
       FOR #tempLoop := 0 TO #NUM_TYPES DO
           //calculate max # of pages
           #recipeMaxPages[#tempLoop] := DINT_TO_INT(CEIL((#tempSetptsUpper[#tempLoop] - #tempSetptsLower[#tempLoop] + 1.0) / #SETPOINTS_PERPAGE));
           //ensure that current page is within the limits
           #recipeCurrentPages[#tempLoop] := LIMIT(MN := 1, IN := #recipeCurrentPages[#tempLoop], MX := #recipeMaxPages[#tempLoop]);
       END_FOR;

       #recipeMaxPages[4] := DINT_TO_INT(CEIL((#tempNumRecipesUpper - #tempNumRecipesLower + 1.0) / #RECIPES_PERPAGE));
       #recipeCurrentPages[4] := LIMIT(MN := 1, IN := #recipeCurrentPages[4], MX := #recipeMaxPages[4]);
   END_REGION


   REGION REAL
       //index in Setpoints_XXX of the current popup
       #tempCurrentPopup := #recipePopupTrackers[#INDEX_REAL] + #SETPOINTS_PERPAGE * (#recipeCurrentPages[#INDEX_REAL] - 1) + #tempSetptsLower[#INDEX_REAL];

       IF #statPrevPopupTrackers[#INDEX_REAL] <> #recipePopupTrackers[#INDEX_REAL] THEN
           //if a new popup has been loaded, load the new setpoint so they can be displayed
           #recipePopup_REAL := #setpoints_REAL[#tempCurrentPopup];
       ELSE
           //if the HMI popup was updated, relay the commands back to the actual setpoint tag for processing
           //taking care to ensure that changes to the setpoints tags made in other areas of the program do not get overwritten
           IF (#statPrevPopupIN_REAL <> #recipePopup_REAL.IN) AND (#statPrevSetpointIN_REAL = #setpoints_REAL[#tempCurrentPopup].IN) THEN
               #setpoints_REAL[#tempCurrentPopup].IN := #recipePopup_REAL.IN;
           END_IF;
           IF #statPrevPopupsSave[#INDEX_REAL] <> #recipePopup_REAL.SaveSetpoint THEN
               #setpoints_REAL[#tempCurrentPopup].SaveSetpoint := #recipePopup_REAL.SaveSetpoint;
           END_IF;
           IF #statPrevPopupsRevert[#INDEX_REAL] <> #recipePopup_REAL.RevertSetpoint THEN
               #setpoints_REAL[#tempCurrentPopup].RevertSetpoint := #recipePopup_REAL.RevertSetpoint;
           END_IF;

           //then update the popup with the latest setpoint information
           #recipePopup_REAL := #setpoints_REAL[#tempCurrentPopup];
       END_IF;

       //set previous values for next scan
       #statPrevPopupIN_REAL := #recipePopup_REAL.IN;
       #statPrevSetpointIN_REAL := #setpoints_REAL[#tempCurrentPopup].IN;
       #statPrevPopupsSave[#INDEX_REAL] := #recipePopup_REAL.SaveSetpoint;
       #statPrevPopupsRevert[#INDEX_REAL] := #recipePopup_REAL.RevertSetpoint;


       //update main setpoint display with setpoint data
       FOR #tempLoop := 0 TO #SETPOINTS_PERPAGE - 1 DO
           IF #tempLoop + #SETPOINTS_PERPAGE * (#recipeCurrentPages[#INDEX_REAL] - 1) + #tempSetptsLower[#INDEX_REAL] <= #tempSetptsUpper[#INDEX_REAL] THEN
               #setpointsArray_REAL[#tempLoop] := #setpoints_REAL[#tempLoop + #SETPOINTS_PERPAGE * (#recipeCurrentPages[#INDEX_REAL] - 1) + #tempSetptsLower[#INDEX_REAL]];
               #setpointFaceplatesDisable_REAL[#tempLoop] := false;
           ELSE
               #setpointFaceplatesDisable_REAL[#tempLoop] := true;
           END_IF;
       END_FOR;
   END_REGION


   REGION DINT
       //index in Setpoints_XXX of the current popup
       #tempCurrentPopup := #recipePopupTrackers[#INDEX_DINT] + #SETPOINTS_PERPAGE * (#recipeCurrentPages[#INDEX_DINT] - 1) + #tempSetptsLower[#INDEX_DINT];

       IF #statPrevPopupTrackers[#INDEX_DINT] <> #recipePopupTrackers[#INDEX_DINT] THEN
           //if a new popup has been loaded, load the new setpoint so they can be displayed
           #recipePopup_DINT := #setpoints_DINT[#tempCurrentPopup];
       ELSE
           //if the HMI popup was updated, relay the commands back to the actual setpoint tag for processing
           //taking care to ensure that changes to the setpoints tags made in other areas of the program do not get overwritten
           IF (#statPrevPopupIN_DINT <> #recipePopup_DINT.IN) AND (#statPrevSetpointIN_DINT = #setpoints_DINT[#tempCurrentPopup].IN) THEN
               #setpoints_DINT[#tempCurrentPopup].IN := #recipePopup_DINT.IN;
           END_IF;
           IF #statPrevPopupsSave[#INDEX_DINT] <> #recipePopup_DINT.SaveSetpoint THEN
               #setpoints_DINT[#tempCurrentPopup].SaveSetpoint := #recipePopup_DINT.SaveSetpoint;
           END_IF;
           IF #statPrevPopupsRevert[#INDEX_DINT] <> #recipePopup_DINT.RevertSetpoint THEN
               #setpoints_DINT[#tempCurrentPopup].RevertSetpoint := #recipePopup_DINT.RevertSetpoint;
           END_IF;

           //then update the popup with the latest setpoint information
           #recipePopup_DINT := #setpoints_DINT[#tempCurrentPopup];
       END_IF;

       //set previous values for next scan
       #statPrevPopupIN_DINT := #recipePopup_DINT.IN;
       #statPrevSetpointIN_DINT := #setpoints_DINT[#tempCurrentPopup].IN;
       #statPrevPopupsSave[#INDEX_DINT] := #recipePopup_DINT.SaveSetpoint;
       #statPrevPopupsRevert[#INDEX_DINT] := #recipePopup_DINT.RevertSetpoint;


       //update main setpoint display with setpoint data
       FOR #tempLoop :=  0 TO #SETPOINTS_PERPAGE - 1 DO
           IF #tempLoop + #SETPOINTS_PERPAGE * (#recipeCurrentPages[#INDEX_DINT] - 1) + #tempSetptsLower[#INDEX_DINT] <= #tempSetptsUpper[#INDEX_DINT] THEN
               #setpointsArray_DINT[#tempLoop] := #setpoints_DINT[#tempLoop + #SETPOINTS_PERPAGE * (#recipeCurrentPages[#INDEX_DINT] - 1) + #tempSetptsLower[#INDEX_DINT]];
               #"setpoint FaceplatesDisable_DINT"[#tempLoop] := false;
           ELSE
               #"setpoint FaceplatesDisable_DINT"[#tempLoop] := true;
           END_IF;
       END_FOR;
   END_REGION


   REGION BOOL
       //index in Setpoints_XXX of the current popup
       #tempCurrentPopup := #recipePopupTrackers[#INDEX_BOOL] + #SETPOINTS_PERPAGE * (#recipeCurrentPages[#INDEX_BOOL] - 1) + #tempSetptsLower[#INDEX_BOOL];

       IF #statPrevPopupTrackers[#INDEX_BOOL] <> #recipePopupTrackers[#INDEX_BOOL] THEN
           //if a new popup has been loaded, load the new setpoint so they can be displayed
           #recipePopup_BOOL := #setpoints_BOOL[#tempCurrentPopup];
       ELSE
           //if the HMI popup was updated, relay the commands back to the actual setpoint tag for processing
           //taking care to ensure that changes to the setpoints tags made in other areas of the program do not get overwritten
           IF (#statPrevPopupIn_BOOL <> #recipePopup_BOOL.IN) AND (#statPrevSetpointIn_BOOL = #setpoints_BOOL[#tempCurrentPopup].IN) THEN
               #setpoints_BOOL[#tempCurrentPopup].IN := #recipePopup_BOOL.IN;
           END_IF;
           IF #statPrevPopupsSave[#INDEX_BOOL] <> #recipePopup_BOOL.SaveSetpoint THEN
               #setpoints_BOOL[#tempCurrentPopup].SaveSetpoint := #recipePopup_BOOL.SaveSetpoint;
           END_IF;
           IF #statPrevPopupsRevert[#INDEX_BOOL] <> #recipePopup_BOOL.RevertSetpoint THEN
               #setpoints_BOOL[#tempCurrentPopup].RevertSetpoint := #recipePopup_BOOL.RevertSetpoint;
           END_IF;

           //then update the popup with the latest setpoint information
           #recipePopup_BOOL := #setpoints_BOOL[#tempCurrentPopup];
       END_IF;

       //set previous values for next scan
       #statPrevPopupIn_BOOL := #recipePopup_BOOL.IN;
       #statPrevSetpointIn_BOOL := #setpoints_BOOL[#tempCurrentPopup].IN;
       #statPrevPopupsSave[#INDEX_BOOL] := #recipePopup_BOOL.SaveSetpoint;
       #statPrevPopupsRevert[#INDEX_BOOL] := #recipePopup_BOOL.RevertSetpoint;


       //update main setpoint display with setpoint data
       FOR #tempLoop := 0 TO #SETPOINTS_PERPAGE-1 DO
           IF #tempLoop + #SETPOINTS_PERPAGE * (#recipeCurrentPages[#INDEX_BOOL] - 1) + #tempSetptsLower[#INDEX_BOOL] <= #tempSetptsUpper[#INDEX_BOOL] THEN
               #setpointsArray_BOOL[#tempLoop] := #setpoints_BOOL[#tempLoop + #SETPOINTS_PERPAGE * (#recipeCurrentPages[#INDEX_BOOL] - 1) + #tempSetptsLower[#INDEX_BOOL]];
               #"setpoint FaceplatesDisable_BOOL"[#tempLoop] := false;
           ELSE
               #"setpoint FaceplatesDisable_BOOL"[#tempLoop] := true;
           END_IF;
       END_FOR;
   END_REGION


   REGION STRING
       //index in Setpoints_XXX of the current popup
       #tempCurrentPopup := #recipePopupTrackers[#INDEX_STRING] + #SETPOINTS_PERPAGE * (#recipeCurrentPages[#INDEX_STRING] - 1) + #tempSetptsLower[#INDEX_STRING];

       IF #statPrevPopupTrackers[#INDEX_STRING] <> #recipePopupTrackers[#INDEX_STRING] THEN
           //if a new popup has been loaded, load the new setpoint so they can be displayed
           #recipePopup_STRING := #setpoints_STRING[#tempCurrentPopup];
       ELSE
           //if the HMI popup was updated, relay the commands back to the actual setpoint tag for processing
           //taking care to ensure that changes to the setpoints tags made in other areas of the program do not get overwritten
           IF (#statPrevPopupIn_STRING <> #recipePopup_STRING.IN) AND (#statPrevSetpointIn_STRING = #setpoints_STRING[#tempCurrentPopup].IN) THEN
               #setpoints_STRING[#tempCurrentPopup].IN := #recipePopup_STRING.IN;
           END_IF;
           IF #statPrevPopupsSave[#INDEX_STRING] <> #recipePopup_STRING.SaveSetpoint THEN
               #setpoints_STRING[#tempCurrentPopup].SaveSetpoint := #recipePopup_STRING.SaveSetpoint;
           END_IF;
           IF #statPrevPopupsRevert[#INDEX_STRING] <> #recipePopup_STRING.RevertSetpoint THEN
               #setpoints_STRING[#tempCurrentPopup].RevertSetpoint := #recipePopup_STRING.RevertSetpoint;
           END_IF;

           //then update the popup with the latest setpoint information
           #recipePopup_STRING := #setpoints_STRING[#tempCurrentPopup];
       END_IF;

       //set previous values for next scan
       #statPrevPopupIn_STRING := #recipePopup_STRING.IN;
       #statPrevSetpointIn_STRING := #setpoints_STRING[#tempCurrentPopup].IN;
       #statPrevPopupsSave[#INDEX_STRING] := #recipePopup_STRING.SaveSetpoint;
       #statPrevPopupsRevert[#INDEX_STRING] := #recipePopup_STRING.RevertSetpoint;


       //update main setpoint display with setpoint data
       FOR #tempLoop := 0 TO #SETPOINTS_PERPAGE - 1 DO
           IF #tempLoop + #SETPOINTS_PERPAGE * (#recipeCurrentPages[#INDEX_STRING] - 1) + #tempSetptsLower[#INDEX_STRING] <= #tempSetptsUpper[#INDEX_STRING] THEN
               #setpointsArray_STRING[#tempLoop] := #setpoints_STRING[#tempLoop + #SETPOINTS_PERPAGE * (#recipeCurrentPages[#INDEX_STRING] - 1) + #tempSetptsLower[#INDEX_STRING]];
               #"setpoint FaceplatesDisable_STRING"[#tempLoop] := false;
           ELSE
               #"setpoint FaceplatesDisable_STRING"[#tempLoop] := true;
           END_IF;
       END_FOR;
   END_REGION


   REGION RECIPE NAMES AND TIMES
       //update the recipe arrays, save times, cum times, and numbers with their current values
       //these values are read only so no need to update the "Recipe Names Array" like we did with the popups
       FOR #tempLoop := 0 TO #RECIPES_PERPAGE - 1 DO
           IF #tempLoop + #RECIPES_PERPAGE * (#recipeCurrentPages[4] - 1) + #tempNumRecipesLower <= #tempNumRecipesUpper THEN
               #recipeArrayNames[#tempLoop] := #recipeNamesArray[#tempLoop + #RECIPES_PERPAGE * (#recipeCurrentPages[4] - 1) + #tempNumRecipesLower];
               #recipeArraySaves[#tempLoop] := #recipeSavesArray[#tempLoop + #RECIPES_PERPAGE * (#recipeCurrentPages[4] - 1) + #tempNumRecipesLower];
               #recipeArrayTimes[#tempLoop] := #recipeTimesArray[#tempLoop + #RECIPES_PERPAGE * (#recipeCurrentPages[4] - 1) + #tempNumRecipesLower];
               #recipeArrayNums[#tempLoop] := #tempLoop + #RECIPES_PERPAGE * (#recipeCurrentPages[4] - 1) + #tempNumRecipesLower;
               #recipeArrayDisables[#tempLoop] := false;
           ELSE
               #recipeArrayDisables[#tempLoop] := true;
           END_IF;
       END_FOR;
   END_REGION





   //update previous values
   #statPrevCurrentPages := #recipeCurrentPages;
   #statPrevPopupTrackers := #recipePopupTrackers;

   //  -------------- END OF LOGIC -------------------------
   ENO := TRUE;   // Set the ENO output
END_FUNCTION_BLOCK

FUNCTION_BLOCK "CPG_RecipeSetpoint_BOOL"   // FB31614, SCL
TITLE = CPG_RecipeSetpoint_BOOL
{ S7_Optimized_Access := 'TRUE' }
AUTHOR : tech.team.motioncontrol@siemens.com
FAMILY : CPG
VERSION : 1.1
// Support: tech.team.motioncontrol@siemens.com
   VAR_INPUT
      enable : Bool;   // If true, setpoint changes are permitted
      disableRecipeControl : Bool;   // If true, the setpoint is no longer handled as a recipe
   END_VAR
   VAR_OUTPUT
      out : Bool;   // Currently running recipe value
      changeEnabled : Bool;   // Enable input is true, setpoint can be changed
      recipeControlDisabled : Bool;   // The value is not subject to recipe controls
      changeNotAllowed : Bool;   // Change is not permitted due to machine state
      recipeSetpointDifference : Bool;   // The currently running (out) value and setpoint value are not equal
   END_VAR
   VAR_IN_OUT
      recipeControl : "CPG_typeRecipeControl";   // Recipe control tag
      recipeSetpoint : "CPG_typeRecipeSetpoint_BOOL";   // Recipe setpoint tag
   END_VAR
   VAR
      statFirstScan : Bool := true;
      statPrevChangeNum : Int;
      statPrevSaveNum : Int;
      statPrevCopyNum : Int;
      statPrevDeleteNum : Int;
      statPrevOut : Bool;
      statChangeNotAllowedTimer : TON_TIME;
      statTimerEN : Bool;
   END_VAR
   VAR CONSTANT
      DELAY_TIME : Time := T#3s;
   END_VAR
BEGIN
   //============================================================================================================
   // SIEMENS AG
   // (c)Copyright 2019 All Rights Reserved
   //------------------------------------------------------------------------------------------------------------
   // Library: LCPG
   // Tested with: S7-1500 with FW version V2.1
   // Engineering: TIA Portal V14
   // Restrictions: ---
   // Requirements: S7-1500
   // Functionality: instantiate this once in the program for each recipe setpoint of BOOL
   // Support: tech.team.motioncontrol@siemens.com
   //------------------------------------------------------------------------------------------------------------
   // Change log table:
   // Version       Date               Expert in charge    Changes applied
   //  01.01.00     02.01.2019         KB                  Initial Release
   //============================================================================================================
   // Function : CPG_RecipeSetpoint_BOOL
   //============================================================================================================

   // Language Selection
   #recipeSetpoint.CurrentName := #recipeSetpoint.SetpointName[#recipeControl.LanguageSelection];
   #recipeSetpoint.CurrentTextFalse := #recipeSetpoint.Text_False[#recipeControl.LanguageSelection];
   #recipeSetpoint.CurrentTextTrue := #recipeSetpoint.Text_True[#recipeControl.LanguageSelection];

   //Recipe Disable Control
   #recipeSetpoint.DisableRecipeControl := #disableRecipeControl;

   //Pass through enable bit
   #recipeSetpoint.SetpointChangeEnabled := #enable;

   //Set out value to match initial one on first scan
   IF #statFirstScan THEN
       #recipeSetpoint.CurrentRecipeValue := #recipeSetpoint.RecipeValues[#recipeControl.CurrentRecipeID];
       #recipeSetpoint.OUT := #recipeSetpoint.RecipeValues[#recipeControl.CurrentRecipeID];
       #statFirstScan := false;
   END_IF;


   REGION RECIPE CONTROL
       // Recipe Control - Change, Save, Copy, Delete, Revert setpoint, Save setpoint
       IF NOT (#recipeSetpoint.DisableRecipeControl) THEN
           //Recipe Change Command
           IF #recipeControl.RecipeChangeNum <> #statPrevChangeNum THEN
               #recipeSetpoint.OUT := #recipeSetpoint.RecipeValues[#recipeControl.CurrentRecipeID];
               #statPrevChangeNum := #recipeControl.RecipeChangeNum;
               // Prevents multiple commands from being executed if this instruction is not being scanned
               #statPrevSaveNum := #recipeControl.RecipeSaveNum;
               #statPrevCopyNum := #recipeControl.RecipeCopyNum;
               #statPrevDeleteNum := #recipeControl.RecipeDeleteNum;
           END_IF;
           //Recipe Save Command
           IF #recipeControl.RecipeSaveNum <> #statPrevSaveNum THEN
               #recipeSetpoint.RecipeValues[#recipeControl.RecipeDestinationID] := #recipeSetpoint.OUT;
               #statPrevSaveNum := #recipeControl.RecipeSaveNum;
               // Prevents multiple commands from being executed if this instruction is not being scanned
               #statPrevCopyNum := #recipeControl.RecipeCopyNum;
               #statPrevDeleteNum := #recipeControl.RecipeDeleteNum;
           END_IF;
           //Recipe Copy Command
           IF #recipeControl.RecipeCopyNum <> #statPrevCopyNum THEN
               #recipeSetpoint.RecipeValues[#recipeControl.RecipeDestinationID] := #recipeSetpoint.RecipeValues[#recipeControl.RecipeSourceID];
               #statPrevCopyNum := #recipeControl.RecipeCopyNum;
               // Prevents multiple commands from being executed if this instruction is not being scanned
               #statPrevDeleteNum := #recipeControl.RecipeDeleteNum;
           END_IF;
           //Recipe Delete Command
           IF #recipeControl.RecipeDeleteNum <> #statPrevDeleteNum THEN
               //edit this line to change the value a deleted recipe defaults to
               #recipeSetpoint.RecipeValues[#recipeControl.RecipeDestinationID] := false;
               #statPrevDeleteNum := #recipeControl.RecipeDeleteNum;
           END_IF;
           // Revert setpoint to saved value
           IF #recipeSetpoint.RevertSetpoint THEN
               #recipeSetpoint.OUT := #recipeSetpoint.RecipeValues[#recipeControl.CurrentRecipeID];
           END_IF;
           //Detect recipe/setpoint difference
           IF (#recipeSetpoint.RecipeValues[#recipeControl.CurrentRecipeID] <> #recipeSetpoint.OUT) AND NOT (#recipeControl.RecipeChange) THEN
               #recipeControl.RecipeSetpointDiff := true;  //signal to recipe control that a setpoint differs
               #recipeSetpoint.RecipeSetpointDiff := true;
           ELSE
               #recipeSetpoint.RecipeSetpointDiff := false;
           END_IF;
           //Save setpoint
           IF #recipeSetpoint.SaveSetpoint THEN
               #recipeSetpoint.RecipeValues[#recipeControl.CurrentRecipeID] := #recipeSetpoint.OUT;
           END_IF;

           //update values stored for current recipe & recipes A, B, & C
           #recipeSetpoint.CurrentRecipeValue := #recipeSetpoint.RecipeValues[#recipeControl.CurrentRecipeID];
           #recipeSetpoint.RecipeValueA := #recipeSetpoint.RecipeValues[#recipeControl.RecipeID_A];
           #recipeSetpoint.RecipeValueB := #recipeSetpoint.RecipeValues[#recipeControl.RecipeID_B];
           #recipeSetpoint.RecipeValueC := #recipeSetpoint.RecipeValues[#recipeControl.RecipeID_C];

       ELSE    //if recipe control is disabled, just update counters
           #recipeSetpoint.RecipeSetpointDiff := false;
           #statPrevChangeNum := #recipeControl.RecipeChangeNum;
           #statPrevSaveNum := #recipeControl.RecipeSaveNum;
           #statPrevCopyNum := #recipeControl.RecipeCopyNum;
           #statPrevDeleteNum := #recipeControl.RecipeDeleteNum;
       END_IF;
   END_REGION


   REGION UPDATE IN VALUE
       //If ENABLE, then changes to the setpoint value are possible
       //otherwise, updating the setpoint is not possible via changing RecipeSetpoint.IN
       IF #enable THEN
           //Clear status bit
           #recipeSetpoint.SetpointChangeDisabled := false;

           // Check for input changed (due to user updating RecipeSetpoint.IN)
           IF (#recipeSetpoint.IN XOR #recipeSetpoint.OUT) AND NOT (#recipeSetpoint.OUT XOR #statPrevOut) THEN
               #recipeSetpoint.OUT := #recipeSetpoint.IN;
           ELSE  // otherwise, update in to match out (this branch can execute due to a recipe change)
               #recipeSetpoint.IN := #recipeSetpoint.OUT;
           END_IF;

       ELSE

           // If in changes, revert and display message
           IF (#recipeSetpoint.IN XOR #recipeSetpoint.OUT) OR #recipeSetpoint.RevertSetpoint THEN
               #recipeSetpoint.IN := #recipeSetpoint.OUT;
               #statTimerEN := false;
               #recipeSetpoint.SetpointChangeDisabled := true;
           END_IF;

           //display "setpoint changes not allowed" 3 seconds after inputting an invalid change
           #statChangeNotAllowedTimer(IN := #statTimerEN,
                                  PT := #DELAY_TIME);

           // Continue to display the status bits for the duration of the timer.
           IF #recipeSetpoint.SetpointChangeDisabled THEN
               #statTimerEN := true;
               #recipeSetpoint.SetpointChangeDisabled :=
                   #recipeSetpoint.SetpointChangeDisabled AND #statTimerEN AND NOT #statChangeNotAllowedTimer.Q;
           END_IF;

       END_IF;
   END_REGION


   REGION DETERMINE HMI TEXTS
       //This is a workaround because multiplexing inside a faceplate is not possible in V14SP1
       IF #recipeSetpoint.OUT THEN
           #recipeSetpoint.Out_Text := #recipeSetpoint.CurrentTextTrue;
       ELSE
           #recipeSetpoint.Out_Text := #recipeSetpoint.CurrentTextFalse;
       END_IF;
       IF #recipeSetpoint.CurrentRecipeValue THEN
           #recipeSetpoint.CurrentRecipeValue_Text := #recipeSetpoint.CurrentTextTrue;
       ELSE
           #recipeSetpoint.CurrentRecipeValue_Text := #recipeSetpoint.CurrentTextFalse;
       END_IF;
       IF #recipeSetpoint.RecipeValueA THEN
           #recipeSetpoint.RecipeA_Text := #recipeSetpoint.CurrentTextTrue;
       ELSE
           #recipeSetpoint.RecipeA_Text := #recipeSetpoint.CurrentTextFalse;
       END_IF;
       IF #recipeSetpoint.RecipeValueB THEN
           #recipeSetpoint.RecipeB_Text := #recipeSetpoint.CurrentTextTrue;
       ELSE
           #recipeSetpoint.RecipeB_Text := #recipeSetpoint.CurrentTextFalse;
       END_IF;
       IF #recipeSetpoint.RecipeValueC THEN
           #recipeSetpoint.RecipeC_Text := #recipeSetpoint.CurrentTextTrue;
       ELSE
           #recipeSetpoint.RecipeC_Text := #recipeSetpoint.CurrentTextFalse;
       END_IF;
   END_REGION


   REGION SET OUTPUTS
       #out := #recipeSetpoint.OUT;
       #statPrevOut := #recipeSetpoint.OUT;
       #changeNotAllowed := #recipeSetpoint.SetpointChangeDisabled;
       #recipeSetpointDifference := #recipeSetpoint.RecipeSetpointDiff;
       #recipeControlDisabled := #recipeSetpoint.DisableRecipeControl;
       #changeEnabled := #recipeSetpoint.SetpointChangeEnabled;
   END_REGION


   //  -------------- END OF LOGIC -------------------------
   ENO := TRUE;   // Set the ENO output
END_FUNCTION_BLOCK

FUNCTION_BLOCK "CPG_RecipeSetpoint_DINT"   // FB31615, SCL
TITLE = CPG_RecipeSetpoint_DINT
{ S7_Optimized_Access := 'TRUE' }
AUTHOR : tech.team.motioncontrol@siemens.com
FAMILY : CPG
VERSION : 1.1
// Support: tech.team.motioncontrol@siemens.com
   VAR_INPUT
      enable : Bool;   // If true, setpoint changes are permitted
      disableRecipeControl : Bool;   // If true, the setpoint is no longer handled as a recipe
   END_VAR
   VAR_OUTPUT
      out : Real;   // Currently running recipe value
      changeEnabled : Bool;   // Enable input is true, setpoint can be changed
      recipeControlDisabled : Bool;   // The value is not subject to recipe controls
      changeNotAllowed : Bool;   // Change is not permitted due to machine state
      recipeSetpointDifference : Bool;   // The currently running (out) value and setpoint value are not equal
      minLimitExceeded : Bool;   // Minimum limit exceeded
      maxLimitExceeded : Bool;   // Maximum limit exceeded
   END_VAR
   VAR_IN_OUT
      recipeControl : "CPG_typeRecipeControl";   // Recipe control tag
      recipeSetpoint : "CPG_typeRecipeSetpoint_DINT";   // Recipe setpoint tag
   END_VAR
   VAR
      statFirstScan : Bool := true;
      statPrevChangeNum : Int;
      statPrevSaveNum : Int;
      statPrevCopyNum : Int;
      statPrevDeleteNum : Int;
      statPrevOut : DInt;
      statLimitsTimer : TP_TIME;
      statLimitsTimerEN : Bool;
      statChangeNotAllowedTimer : TON_TIME;
      statTimerEN : Bool;
   END_VAR
   VAR_TEMP
      tempLimit : DInt;
   END_VAR
   VAR CONSTANT
      DELAY_TIME : Time := T#3s;
   END_VAR
BEGIN
   //============================================================================================================
   // SIEMENS AG
   // (c)Copyright 2019 All Rights Reserved
   //------------------------------------------------------------------------------------------------------------
   // Library: LCPG
   // Tested with: S7-1500 with FW version V2.1
   // Engineering: TIA Portal V14
   // Restrictions: ---
   // Requirements: S7-1500
   // Functionality: instantiate this once in the program for each recipe setpoint of DINT
   // Support: tech.team.motioncontrol@siemens.com
   //------------------------------------------------------------------------------------------------------------
   // Change log table:
   // Version       Date               Expert in charge    Changes applied
   //  01.01.00     02.01.2019         KB                  Initial Release
   //============================================================================================================
   // Function : CPG_RecipeSetpoint_DINT
   //============================================================================================================

   // Language Selection
   #recipeSetpoint.CurrentName := #recipeSetpoint.SetpointName[#recipeControl.LanguageSelection];

   //Recipe Disable Control
   #recipeSetpoint.DisableRecipeControl := #disableRecipeControl;

   //Pass through enable bit
   #recipeSetpoint.SetpointChangeEnabled := #enable;

   //Set out value to match initial one on first scan
   IF #statFirstScan THEN
       #recipeSetpoint.CurrentRecipeValue := #recipeSetpoint.RecipeValues[#recipeControl.CurrentRecipeID];
       #recipeSetpoint.OUT := #recipeSetpoint.RecipeValues[#recipeControl.CurrentRecipeID];
       #statFirstScan := false;
   END_IF;


   REGION CHECK LIMITS
       //checks if min & max limits are valid.  If they are not in order, swap them
       IF #recipeSetpoint.minLimit > #recipeSetpoint.maxLimit THEN
           #tempLimit := #recipeSetpoint.minLimit;
           #recipeSetpoint.minLimit := #recipeSetpoint.maxLimit;
           #recipeSetpoint.maxLimit := #tempLimit;
       END_IF;

       //checks if the saved recipe value is outside the bounds, either due to a runtime change of the limits or a bad configuration
       //if problems, and recipe control is on, set the saved value to the default (min limit, same as recipeDelete)
       //Note that this check is only on the current recipe, and also is only performed if recipeControlDisable is false
       IF #recipeSetpoint.RecipeValues[#recipeControl.CurrentRecipeID] < #recipeSetpoint.minLimit
           OR #recipeSetpoint.RecipeValues[#recipeControl.CurrentRecipeID] > #recipeSetpoint.maxLimit
           AND NOT (#recipeSetpoint.DisableRecipeControl) THEN
           #recipeSetpoint.RecipeValues[#recipeControl.CurrentRecipeID] := #recipeSetpoint.minLimit;
       END_IF;

       //Checks the out value.  Note that this value matters even if recipeControlDisable is true
       //If the value is a being controlled, then set the value to the (guarenteed to be in range) saved recipe value
       //If the value is not being treated as a recipe, set it to the default (minlimit)
       IF #recipeSetpoint.OUT < #recipeSetpoint.minLimit OR #recipeSetpoint.OUT > #recipeSetpoint.maxLimit THEN
           IF NOT (#recipeSetpoint.DisableRecipeControl) THEN
               #recipeSetpoint.OUT := #recipeSetpoint.RecipeValues[#recipeControl.CurrentRecipeID];
           ELSE
               #recipeSetpoint.OUT := #recipeSetpoint.minLimit;
           END_IF;
       END_IF;
   END_REGION


   REGION RECIPE CONTROL
       // Recipe Control - Change, Save, Copy, Delete, Revert setpoint, Save setpoint
       IF NOT (#recipeSetpoint.DisableRecipeControl) THEN
           //Recipe Change Command
           IF #recipeControl.RecipeChangeNum <> #statPrevChangeNum THEN
               #recipeSetpoint.OUT := #recipeSetpoint.RecipeValues[#recipeControl.CurrentRecipeID];
               #statPrevChangeNum := #recipeControl.RecipeChangeNum;
               // Prevents multiple commands from being executed if this instruction is not being scanned
               #statPrevSaveNum := #recipeControl.RecipeSaveNum;
               #statPrevCopyNum := #recipeControl.RecipeCopyNum;
               #statPrevDeleteNum := #recipeControl.RecipeDeleteNum;
           END_IF;
           //Recipe Save Command
           IF #recipeControl.RecipeSaveNum <> #statPrevSaveNum THEN
               #recipeSetpoint.RecipeValues[#recipeControl.RecipeDestinationID] := #recipeSetpoint.OUT;
               #statPrevSaveNum := #recipeControl.RecipeSaveNum;
               // Prevents multiple commands from being executed if this instruction is not being scanned
               #statPrevCopyNum := #recipeControl.RecipeCopyNum;
               #statPrevDeleteNum := #recipeControl.RecipeDeleteNum;
           END_IF;
           //Recipe Copy Command
           IF #recipeControl.RecipeCopyNum <> #statPrevCopyNum THEN
               #recipeSetpoint.RecipeValues[#recipeControl.RecipeDestinationID] := #recipeSetpoint.RecipeValues[#recipeControl.RecipeSourceID];
               #statPrevCopyNum := #recipeControl.RecipeCopyNum;
               // Prevents multiple commands from being executed if this instruction is not being scanned
               #statPrevDeleteNum := #recipeControl.RecipeDeleteNum;
           END_IF;
           //Recipe Delete Command
           IF #recipeControl.RecipeDeleteNum <> #statPrevDeleteNum THEN
               //edit this line to change the value a deleted recipe defaults to
               #recipeSetpoint.RecipeValues[#recipeControl.RecipeDestinationID] := #recipeSetpoint.minLimit;
               #statPrevDeleteNum := #recipeControl.RecipeDeleteNum;
           END_IF;
           // Revert setpoint to saved value
           IF #recipeSetpoint.RevertSetpoint THEN
               #recipeSetpoint.OUT := #recipeSetpoint.RecipeValues[#recipeControl.CurrentRecipeID];
           END_IF;
           //Detect recipe/setpoint difference
           IF (#recipeSetpoint.RecipeValues[#recipeControl.CurrentRecipeID] <> #recipeSetpoint.OUT) AND NOT (#recipeControl.RecipeChange) THEN
               #recipeControl.RecipeSetpointDiff := true;  //signal to recipe control that a setpoint differs
               #recipeSetpoint.RecipeSetpointDiff := true;
           ELSE
               #recipeSetpoint.RecipeSetpointDiff := false;
           END_IF;
           //Save setpoint
           IF #recipeSetpoint.SaveSetpoint THEN
               #recipeSetpoint.RecipeValues[#recipeControl.CurrentRecipeID] := #recipeSetpoint.OUT;
           END_IF;

           //update values stored for current recipe & recipes A, B, & C
           #recipeSetpoint.CurrentRecipeValue := #recipeSetpoint.RecipeValues[#recipeControl.CurrentRecipeID];
           #recipeSetpoint.RecipeValueA := #recipeSetpoint.RecipeValues[#recipeControl.RecipeID_A];
           #recipeSetpoint.RecipeValueB := #recipeSetpoint.RecipeValues[#recipeControl.RecipeID_B];
           #recipeSetpoint.RecipeValueC := #recipeSetpoint.RecipeValues[#recipeControl.RecipeID_C];

       ELSE    //if recipe control is disabled, just update counters
           #recipeSetpoint.RecipeSetpointDiff := false;
           #statPrevChangeNum := #recipeControl.RecipeChangeNum;
           #statPrevSaveNum := #recipeControl.RecipeSaveNum;
           #statPrevCopyNum := #recipeControl.RecipeCopyNum;
           #statPrevDeleteNum := #recipeControl.RecipeDeleteNum;
       END_IF;
   END_REGION

   REGION UPDATE IN VALUE
       //If ENABLE, then changes to the setpoint value are possible
       //otherwise, updating the setpoint is not possible via changing RecipeSetpoint.IN
       IF #enable THEN
           //Clear status bit
           #recipeSetpoint.SetpointChangeDisabled := false;

           // Check for value within limits and input changed (due to user updating RecipeSetpoint.IN)
           IF (#recipeSetpoint.minLimit <= #recipeSetpoint.IN) AND (#recipeSetpoint.IN <= #recipeSetpoint.maxLimit) AND
               (#recipeSetpoint.IN <> #recipeSetpoint.OUT) AND (#recipeSetpoint.OUT = #statPrevOut) THEN
               #recipeSetpoint.OUT := #recipeSetpoint.IN;
               #recipeSetpoint.minLimitReached := false;
               #recipeSetpoint.maxLimitReached := false;
           // Check for value within limits and output changed (due to a recipe change)
           ELSIF (#recipeSetpoint.minLimit <= #recipeSetpoint.IN) AND (#recipeSetpoint.IN <= #recipeSetpoint.maxLimit) AND
               (#recipeSetpoint.IN <> #recipeSetpoint.OUT) AND (#recipeSetpoint.OUT <> #statPrevOut) THEN
               #recipeSetpoint.IN := #recipeSetpoint.OUT;
               #recipeSetpoint.minLimitReached := false;
               #recipeSetpoint.maxLimitReached := false;
           // Check for value below minimum limit
           ELSIF (#recipeSetpoint.minLimit > #recipeSetpoint.IN) THEN
               #statLimitsTimerEN := true;
               #recipeSetpoint.IN := #recipeSetpoint.OUT;
               #recipeSetpoint.minLimitReached := true;
               #recipeSetpoint.maxLimitReached := false;
           // Check for value above maximum limit
           ELSIF (#recipeSetpoint.maxLimit < #recipeSetpoint.IN) THEN
               #statLimitsTimerEN := true;
               #recipeSetpoint.IN := #recipeSetpoint.OUT;
               #recipeSetpoint.minLimitReached := false;
               #recipeSetpoint.maxLimitReached := true;
           END_IF;

           #statLimitsTimer(IN := #statLimitsTimerEN,
                        PT := #DELAY_TIME);

           // Continue to display the status bits for the duration of the timer.
           IF #recipeSetpoint.minLimitReached OR #recipeSetpoint.maxLimitReached THEN
               #statLimitsTimerEN := false;
               #recipeSetpoint.minLimitReached := #recipeSetpoint.minLimitReached AND #statLimitsTimer.Q;
               #recipeSetpoint.maxLimitReached := #recipeSetpoint.maxLimitReached AND #statLimitsTimer.Q;
           END_IF;

       ELSE

           // If IN changes, revert and display message
           IF (#recipeSetpoint.IN <> #recipeSetpoint.OUT) OR #recipeSetpoint.RevertSetpoint THEN
               #recipeSetpoint.IN := #recipeSetpoint.OUT;
               #statTimerEN := false;
               #recipeSetpoint.SetpointChangeDisabled := true;
               #recipeSetpoint.minLimitReached := false;
               #recipeSetpoint.maxLimitReached := false;
           END_IF;

           //display "setpoint changes not allowed" 3 seconds after inputting an invalid change
           #statChangeNotAllowedTimer(IN := #statTimerEN,
                                  PT := #DELAY_TIME);

           // Continue to display the status bits for the duration of the timer.
           IF #recipeSetpoint.SetpointChangeDisabled THEN
               #statTimerEN := true;
               #recipeSetpoint.SetpointChangeDisabled :=
                   #recipeSetpoint.SetpointChangeDisabled AND #statTimerEN AND NOT #statChangeNotAllowedTimer.Q;
           END_IF;

       END_IF;
   END_REGION


   REGION SET OUTPUTS
       #out := #recipeSetpoint.OUT;
       #statPrevOut := #recipeSetpoint.OUT;
       #changeNotAllowed := #recipeSetpoint.SetpointChangeDisabled;
       #recipeSetpointDifference := #recipeSetpoint.RecipeSetpointDiff;
       #recipeControlDisabled := #recipeSetpoint.DisableRecipeControl;
       #changeEnabled := #recipeSetpoint.SetpointChangeEnabled;
       #minLimitExceeded := #recipeSetpoint.minLimitReached;
       #maxLimitExceeded := #recipeSetpoint.maxLimitReached;
   END_REGION

   //  -------------- END OF LOGIC -------------------------
   ENO := TRUE;   // Set the ENO output
END_FUNCTION_BLOCK

FUNCTION_BLOCK "CPG_RecipeSetpoint_REAL"   // FB31616, SCL
TITLE = CPG_RecipeSetpoint_REAL
{ S7_Optimized_Access := 'TRUE' }
AUTHOR : tech.team.motioncontrol@siemens.com
FAMILY : CPG
VERSION : 1.1
// Support: tech.team.motioncontrol@siemens.com
   VAR_INPUT
      enable : Bool;   // If true, setpoint changes are permitted
      disableRecipeControl : Bool;   // If true, the setpoint is no longer handled as a recipe
   END_VAR
   VAR_OUTPUT
      out : Real;   // Currently running recipe value
      changeEnabled : Bool;   // Enable input is true, setpoint can be changed
      recipeControlDisabled : Bool;   // The value is not subject to recipe controls
      changeNotAllowed : Bool;   // Change is not permitted due to machine state
      recipeSetpointDifference : Bool;   // The currently running (out) value and setpoint value are not equal
      minLimitExceeded : Bool;   // Minimum limit exceeded
      maxLimitExceeded : Bool;   // Maximum limit exceeded
   END_VAR
   VAR_IN_OUT
      recipeControl : "CPG_typeRecipeControl";   // Recipe control tag
      recipeSetpoint : "CPG_typeRecipeSetpoint_REAL";   // Recipe setpoint tag
   END_VAR
   VAR
      statFirstScan : Bool := true;
      statPrevChangeNum : Int;
      statPrevSaveNum : Int;
      statPrevCopyNum : Int;
      statPrevDeleteNum : Int;
      statPrevOut : Real;
      statLimitsTimer : TP_TIME;
      statLimitsTimerEN : Bool;
      statChangeNotAllowedTimer : TON_TIME;
      statTimerEN : Bool;
   END_VAR
   VAR_TEMP
      tempLimit : Real;
   END_VAR
   VAR CONSTANT
      DELAY_TIME : Time := T#3s;
   END_VAR
BEGIN
   //============================================================================================================
   // SIEMENS AG
   // (c)Copyright 2019 All Rights Reserved
   //------------------------------------------------------------------------------------------------------------
   // Library: LCPG
   // Tested with: S7-1500 with FW version V2.1
   // Engineering: TIA Portal V14
   // Restrictions: ---
   // Requirements: S7-1500
   // Functionality: instantiate this once in the program for each recipe setpoint of REAL
   // Support: tech.team.motioncontrol@siemens.com
   //------------------------------------------------------------------------------------------------------------
   // Change log table:
   // Version       Date               Expert in charge    Changes applied
   //  01.01.00     02.01.2019         KB                  Initial Release
   //============================================================================================================
   // Function : CPG_RecipeSetpoint_REAL
   //============================================================================================================

   // Language Selection
   #recipeSetpoint.CurrentName := #recipeSetpoint.SetpointName[#recipeControl.LanguageSelection];

   //Recipe Disable Control
   #recipeSetpoint.DisableRecipeControl := #disableRecipeControl;

   //Pass through enable bit
   #recipeSetpoint.SetpointChangeEnabled := #enable;

   //Set out value to match initial one on first scan
   IF #statFirstScan THEN
       #recipeSetpoint.CurrentRecipeValue := #recipeSetpoint.RecipeValues[#recipeControl.CurrentRecipeID];
       #recipeSetpoint.OUT := #recipeSetpoint.RecipeValues[#recipeControl.CurrentRecipeID];
       #statFirstScan := false;
   END_IF;


   REGION CHECK LIMITS
       //checks if min & max limits are valid.  If they are not in order, swap them
       IF #recipeSetpoint.minLimit > #recipeSetpoint.maxLimit THEN
           #tempLimit := #recipeSetpoint.minLimit;
           #recipeSetpoint.minLimit := #recipeSetpoint.maxLimit;
           #recipeSetpoint.maxLimit := #tempLimit;
       END_IF;

       //checks if the saved recipe value is outside the bounds, either due to a runtime change of the limits or a bad configuration
       //if problems, and recipe control is on, set the saved value to the default (min limit, same as recipeDelete)
       //Note that this check is only on the current recipe, and also is only performed if recipeControlDisable is false
       IF #recipeSetpoint.RecipeValues[#recipeControl.CurrentRecipeID] < #recipeSetpoint.minLimit
           OR #recipeSetpoint.RecipeValues[#recipeControl.CurrentRecipeID] > #recipeSetpoint.maxLimit
           AND NOT (#recipeSetpoint.DisableRecipeControl) THEN
           #recipeSetpoint.RecipeValues[#recipeControl.CurrentRecipeID] := #recipeSetpoint.minLimit;
       END_IF;

       //Checks the out value.  Note that this value matters even if recipeControlDisable is true
       //If the value is a being controlled, then set the value to the (guarenteed to be in range) saved recipe value
       //If the value is not being treated as a recipe, set it to the default (minlimit)
       IF #recipeSetpoint.OUT < #recipeSetpoint.minLimit OR #recipeSetpoint.OUT > #recipeSetpoint.maxLimit THEN
           IF NOT (#recipeSetpoint.DisableRecipeControl) THEN
               #recipeSetpoint.OUT := #recipeSetpoint.RecipeValues[#recipeControl.CurrentRecipeID];
           ELSE
               #recipeSetpoint.OUT := #recipeSetpoint.minLimit;
           END_IF;
       END_IF;
   END_REGION


   REGION RECIPE CONTROL
       // Recipe Control - Change, Save, Copy, Delete, Revert setpoint, Save setpoint
       IF NOT (#recipeSetpoint.DisableRecipeControl) THEN
           //Recipe Change Command
           IF #recipeControl.RecipeChangeNum <> #statPrevChangeNum THEN
               #recipeSetpoint.OUT := #recipeSetpoint.RecipeValues[#recipeControl.CurrentRecipeID];
               #statPrevChangeNum := #recipeControl.RecipeChangeNum;
               // Prevents multiple commands from being executed if this instruction is not being scanned
               #statPrevSaveNum := #recipeControl.RecipeSaveNum;
               #statPrevCopyNum := #recipeControl.RecipeCopyNum;
               #statPrevDeleteNum := #recipeControl.RecipeDeleteNum;
           END_IF;
           //Recipe Save Command
           IF #recipeControl.RecipeSaveNum <> #statPrevSaveNum THEN
               #recipeSetpoint.RecipeValues[#recipeControl.RecipeDestinationID] := #recipeSetpoint.OUT;
               #statPrevSaveNum := #recipeControl.RecipeSaveNum;
               // Prevents multiple commands from being executed if this instruction is not being scanned
               #statPrevCopyNum := #recipeControl.RecipeCopyNum;
               #statPrevDeleteNum := #recipeControl.RecipeDeleteNum;
           END_IF;
           //Recipe Copy Command
           IF #recipeControl.RecipeCopyNum <> #statPrevCopyNum THEN
               #recipeSetpoint.RecipeValues[#recipeControl.RecipeDestinationID] := #recipeSetpoint.RecipeValues[#recipeControl.RecipeSourceID];
               #statPrevCopyNum := #recipeControl.RecipeCopyNum;
               // Prevents multiple commands from being executed if this instruction is not being scanned
               #statPrevDeleteNum := #recipeControl.RecipeDeleteNum;
           END_IF;
           //Recipe Delete Command
           IF #recipeControl.RecipeDeleteNum <> #statPrevDeleteNum THEN
               //edit this line to change the value a deleted recipe defaults to
               #recipeSetpoint.RecipeValues[#recipeControl.RecipeDestinationID] := #recipeSetpoint.minLimit;   
               #statPrevDeleteNum := #recipeControl.RecipeDeleteNum;
           END_IF;
           // Revert setpoint to saved value
           IF #recipeSetpoint.RevertSetpoint THEN
               #recipeSetpoint.OUT := #recipeSetpoint.RecipeValues[#recipeControl.CurrentRecipeID];
           END_IF;
           //Detect recipe/setpoint difference
           IF (#recipeSetpoint.RecipeValues[#recipeControl.CurrentRecipeID] <> #recipeSetpoint.OUT) AND NOT (#recipeControl.RecipeChange) THEN
               #recipeControl.RecipeSetpointDiff := true;  //signal to recipe control that a setpoint differs
               #recipeSetpoint.RecipeSetpointDiff := true;
           ELSE
               #recipeSetpoint.RecipeSetpointDiff := false;
           END_IF;
           //Save setpoint
           IF #recipeSetpoint.SaveSetpoint THEN
               #recipeSetpoint.RecipeValues[#recipeControl.CurrentRecipeID] := #recipeSetpoint.OUT;
           END_IF;


           //update values stored for current recipe & recipes A, B, & C
           #recipeSetpoint.CurrentRecipeValue := #recipeSetpoint.RecipeValues[#recipeControl.CurrentRecipeID];
           #recipeSetpoint.RecipeValueA := #recipeSetpoint.RecipeValues[#recipeControl.RecipeID_A];
           #recipeSetpoint.RecipeValueB := #recipeSetpoint.RecipeValues[#recipeControl.RecipeID_B];
           #recipeSetpoint.RecipeValueC := #recipeSetpoint.RecipeValues[#recipeControl.RecipeID_C];

       ELSE    //if recipe control is disabled, just update counters
           #recipeSetpoint.RecipeSetpointDiff := false;
           #statPrevChangeNum := #recipeControl.RecipeChangeNum;
           #statPrevSaveNum := #recipeControl.RecipeSaveNum;
           #statPrevCopyNum := #recipeControl.RecipeCopyNum;
           #statPrevDeleteNum := #recipeControl.RecipeDeleteNum;
       END_IF;
   END_REGION


   REGION UPDATE IN VALUE
       //If ENABLE, then changes to the setpoint value are possible
       //otherwise, updating the setpoint is not possible via changing RecipeSetpoint.IN
       IF #enable THEN
           //Clear status bit
           #recipeSetpoint.SetpointChangeDisabled := false;

           // Check for value within limits and input changed (due to user updating RecipeSetpoint.IN)
           IF (#recipeSetpoint.minLimit <= #recipeSetpoint.IN) AND (#recipeSetpoint.IN <= #recipeSetpoint.maxLimit) AND
               (#recipeSetpoint.IN <> #recipeSetpoint.OUT) AND (#recipeSetpoint.OUT = #statPrevOut) THEN
               #recipeSetpoint.OUT := #recipeSetpoint.IN;
               #recipeSetpoint.minLimitReached := false;
               #recipeSetpoint.maxLimitReached := false;
           // Check for value within limits and output changed (due to a recipe change)
           ELSIF (#recipeSetpoint.minLimit <= #recipeSetpoint.IN) AND (#recipeSetpoint.IN <= #recipeSetpoint.maxLimit) AND
               (#recipeSetpoint.IN <> #recipeSetpoint.OUT) AND (#recipeSetpoint.OUT <> #statPrevOut) THEN
               #recipeSetpoint.IN := #recipeSetpoint.OUT;
               #recipeSetpoint.minLimitReached := false;
               #recipeSetpoint.maxLimitReached := false;
           // Check for value below minimum limit
           ELSIF (#recipeSetpoint.minLimit > #recipeSetpoint.IN) THEN
               #statLimitsTimerEN := true;
               #recipeSetpoint.IN := #recipeSetpoint.OUT;
               #recipeSetpoint.minLimitReached := true;
               #recipeSetpoint.maxLimitReached := false;
           // Check for value above maximum limit
           ELSIF (#recipeSetpoint.maxLimit < #recipeSetpoint.IN) THEN
               #statLimitsTimerEN := true;
               #recipeSetpoint.IN := #recipeSetpoint.OUT;
               #recipeSetpoint.minLimitReached := false;
               #recipeSetpoint.maxLimitReached := true;
           END_IF;

           #statLimitsTimer(IN := #statLimitsTimerEN,
                        PT := #DELAY_TIME);

           // Continue to display the status bits for the duration of the timer.
           IF #recipeSetpoint.minLimitReached OR #recipeSetpoint.maxLimitReached THEN
               #statLimitsTimerEN := false;
               #recipeSetpoint.minLimitReached := #recipeSetpoint.minLimitReached AND #statLimitsTimer.Q;
               #recipeSetpoint.maxLimitReached := #recipeSetpoint.maxLimitReached AND #statLimitsTimer.Q;
           END_IF;

       ELSE

           // If IN changes, revert and display message
           IF (#recipeSetpoint.IN <> #recipeSetpoint.OUT) OR #recipeSetpoint.RevertSetpoint THEN
               #recipeSetpoint.IN := #recipeSetpoint.OUT;
               #statTimerEN := false;
               #recipeSetpoint.SetpointChangeDisabled := true;
               #recipeSetpoint.minLimitReached := false;
               #recipeSetpoint.maxLimitReached := false;
           END_IF;

           //display "setpoint changes not allowed" 3 seconds after inputting an invalid change
           #statChangeNotAllowedTimer(IN := #statTimerEN,
                                  PT := #DELAY_TIME);

           // Continue to display the status bits for the duration of the timer.
           IF #recipeSetpoint.SetpointChangeDisabled THEN
               #statTimerEN := true;
               #recipeSetpoint.SetpointChangeDisabled :=
                   #recipeSetpoint.SetpointChangeDisabled AND #statTimerEN AND NOT #statChangeNotAllowedTimer.Q;
           END_IF;

       END_IF;
   END_REGION


   REGION SET OUTPUTS
       #out := #recipeSetpoint.OUT;
       #statPrevOut := #recipeSetpoint.OUT;
       #changeNotAllowed := #recipeSetpoint.SetpointChangeDisabled;
       #recipeSetpointDifference := #recipeSetpoint.RecipeSetpointDiff;
       #recipeControlDisabled := #recipeSetpoint.DisableRecipeControl;
       #changeEnabled := #recipeSetpoint.SetpointChangeEnabled;
       #minLimitExceeded := #recipeSetpoint.minLimitReached;
       #maxLimitExceeded := #recipeSetpoint.maxLimitReached;
   END_REGION

   //  -------------- END OF LOGIC -------------------------
   ENO := TRUE;   // Set the ENO output
END_FUNCTION_BLOCK

